REGION Network 2
   // **********************************************************************************************************************
   // 
   // Carrier 81 I-Device Data Transfer Interlocks from Carrier to SDC
   // 
   // **********************************************************************************************************************
   RUNG wire#powerrail
      Coil( "SectionComment" )
   END_RUNG
   // the same network as SCL:
   "SectionComment" := TRUE;
END_REGION

REGION Network 3
   RUNG wire#powerrail
      Contact( "Carrier_81_Status.0" )
      Coil( "EMS".Carrier[81].SDC_IN.HeartBeat )
   END_RUNG
   // the same network as SCL:
   "EMS".Carrier[81].SDC_IN.HeartBeat := "Carrier_81_Status.0";
END_REGION

REGION Network 4
   "C81_Heartbeat_On_Timer".TON(IN := "EMS".Carrier[81].SDC_IN.HeartBeat, PT := T#3s);
END_REGION

REGION Network 5
   "C81_Heartbeat_Off_Timer".TON(IN := NOT "EMS".Carrier[81].SDC_IN.HeartBeat, PT := T#3s);
END_REGION

REGION Network 6
   RUNG wire#powerrail
      Contact( "Carrier_81_Status.7" )
      wire#w1
      Coil( "EMS".Carrier[81].CommFlt )
   END_RUNG
   RUNG wire#powerrail
      Contact( "C81_Heartbeat_On_Timer".Q )
   END_RUNG wire#w1
   RUNG wire#powerrail
      Contact( "C81_Heartbeat_Off_Timer".Q )
   END_RUNG wire#w1
   // the same network as SCL:
   "EMS".Carrier[81].CommFlt := "Carrier_81_Status.7" OR "C81_Heartbeat_On_Timer".Q OR "C81_Heartbeat_Off_Timer".Q;
END_REGION

REGION Network 7
   RUNG wire#powerrail
      Contact( "EMS".Carrier[81].CommFlt )
      JumpCoil( C81_Comm_Fault )
   END_RUNG
   // the same network as SCL:
   IF "EMS".Carrier[81].CommFlt THEN GOTO C81_Comm_Fault; END_IF;
END_REGION

REGION Network 8
   RUNG wire#powerrail
      { S7_Templates := "SrcType := Word" } NE_Contact(in1 := "Carrier_81_CarrierNumber", in2 := 0)
      Move(in := "Carrier_81_CarrierNumber", out1 => "EMS".Carrier[81].SDC_IN.CarrierNumber)
   END_RUNG
   // the same network as SCL:
   IF "Carrier_81_CarrierNumber" <> 0 THEN
       "EMS".Carrier[81].SDC_IN.CarrierNumber := "Carrier_81_CarrierNumber";
   END_IF;
END_REGION

REGION Network 9
   RUNG wire#powerrail
      { S7_Templates := "SrcType := DWord" } NE_Contact(in1 := "Carrier_81_CarrierPosition", in2 := 0)
      Move(in := "Carrier_81_CarrierPosition", out1 => "EMS".Carrier[81].SDC_IN.CarrierPosition)
   END_RUNG
   // the same network as SCL:
   IF "Carrier_81_CarrierPosition" <> 0 THEN
       "EMS".Carrier[81].SDC_IN.CarrierPosition := "Carrier_81_CarrierPosition";
   END_IF;
END_REGION

REGION Network 10
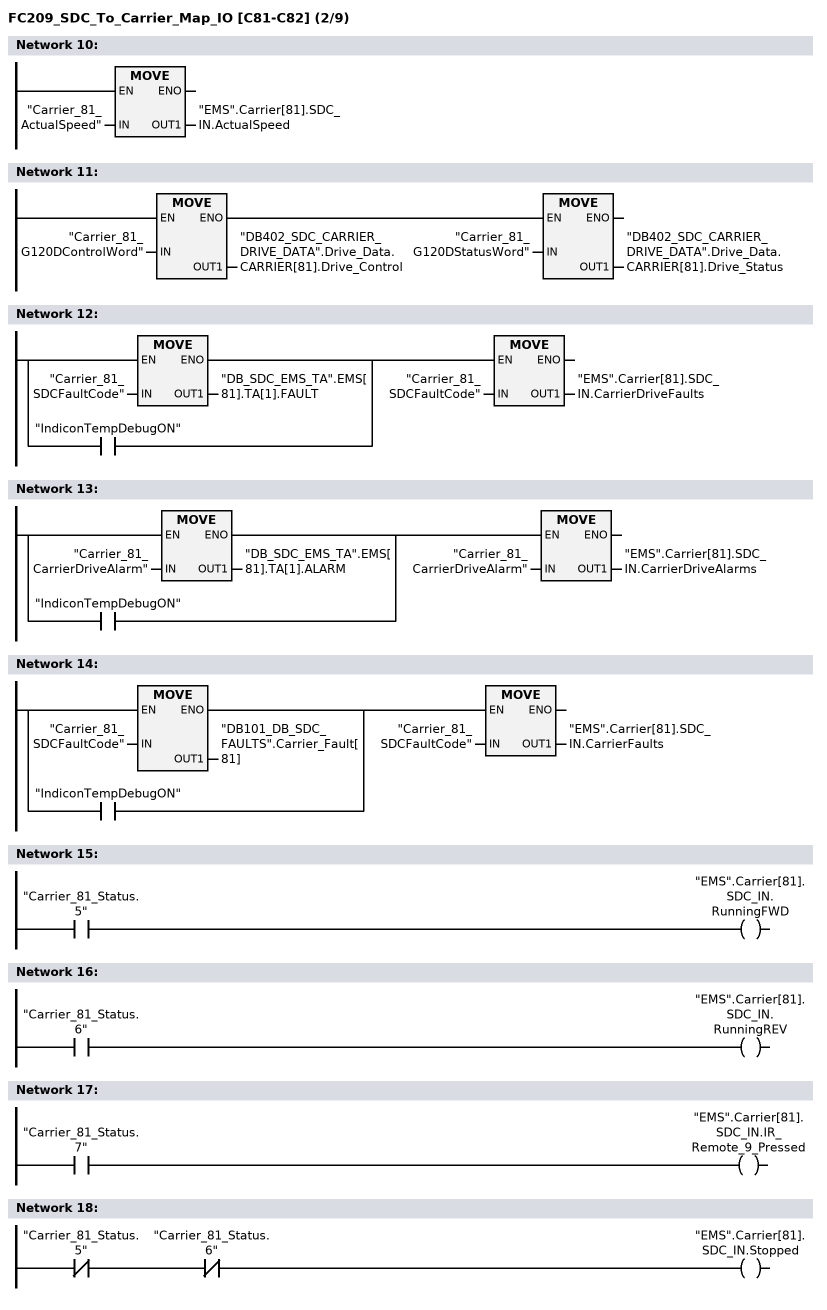
   RUNG wire#powerrail
      Move(in := "Carrier_81_ActualSpeed", out1 => "EMS".Carrier[81].SDC_IN.ActualSpeed)
   END_RUNG
   // the same network as SCL:
   "EMS".Carrier[81].SDC_IN.ActualSpeed := "Carrier_81_ActualSpeed";
END_REGION

REGION Network 11
   RUNG wire#powerrail
      Move(in := "Carrier_81_G120DControlWord", out1 => "DB402_SDC_CARRIER_DRIVE_DATA".Drive_Data.CARRIER[81].Drive_Control)
      Move(in := "Carrier_81_G120DStatusWord", out1 => "DB402_SDC_CARRIER_DRIVE_DATA".Drive_Data.CARRIER[81].Drive_Status)
   END_RUNG
   // the same network as SCL:
   "DB402_SDC_CARRIER_DRIVE_DATA".Drive_Data.CARRIER[81].Drive_Control := "Carrier_81_G120DControlWord";
   "DB402_SDC_CARRIER_DRIVE_DATA".Drive_Data.CARRIER[81].Drive_Status := "Carrier_81_G120DStatusWord";
END_REGION

REGION Network 12
   RUNG wire#powerrail
      Move(in := "Carrier_81_SDCFaultCode", out1 => "DB_SDC_EMS_TA".EMS[81].TA[1].FAULT)
      wire#w1
      Move(in := "Carrier_81_SDCFaultCode", out1 => "EMS".Carrier[81].SDC_IN.CarrierDriveFaults)
   END_RUNG
   RUNG wire#powerrail
      Contact( "IndiconTempDebugON" )
   END_RUNG wire#w1
   // the same network as SCL:
   "DB_SDC_EMS_TA".EMS[81].TA[1].FAULT := "Carrier_81_SDCFaultCode";
   IF TRUE OR "IndiconTempDebugON" THEN
       "EMS".Carrier[81].SDC_IN.CarrierDriveFaults := "Carrier_81_SDCFaultCode";
   END_IF;
END_REGION

REGION Network 13
   RUNG wire#powerrail
      Move(in := "Carrier_81_CarrierDriveAlarm", out1 => "DB_SDC_EMS_TA".EMS[81].TA[1].ALARM)
      wire#w1
      Move(in := "Carrier_81_CarrierDriveAlarm", out1 => "EMS".Carrier[81].SDC_IN.CarrierDriveAlarms)
   END_RUNG
   RUNG wire#powerrail
      Contact( "IndiconTempDebugON" )
   END_RUNG wire#w1
   // the same network as SCL:
   "DB_SDC_EMS_TA".EMS[81].TA[1].ALARM := "Carrier_81_CarrierDriveAlarm";
   IF TRUE OR "IndiconTempDebugON" THEN
       "EMS".Carrier[81].SDC_IN.CarrierDriveAlarms := "Carrier_81_CarrierDriveAlarm";
   END_IF;
END_REGION

REGION Network 14
   RUNG wire#powerrail
      Move(in := "Carrier_81_SDCFaultCode", out1 => "DB101_DB_SDC_FAULTS".Carrier_Fault[81])
      wire#w1
      Move(in := "Carrier_81_SDCFaultCode", out1 => "EMS".Carrier[81].SDC_IN.CarrierFaults)
   END_RUNG
   RUNG wire#powerrail
      Contact( "IndiconTempDebugON" )
   END_RUNG wire#w1
   // the same network as SCL:
   "DB101_DB_SDC_FAULTS".Carrier_Fault[81] := "Carrier_81_SDCFaultCode";
   IF TRUE OR "IndiconTempDebugON" THEN
       "EMS".Carrier[81].SDC_IN.CarrierFaults := "Carrier_81_SDCFaultCode";
   END_IF;
END_REGION

REGION Network 15
   RUNG wire#powerrail
      Contact( "Carrier_81_Status.5" )
      Coil( "EMS".Carrier[81].SDC_IN.RunningFWD )
   END_RUNG
   // the same network as SCL:
   "EMS".Carrier[81].SDC_IN.RunningFWD := "Carrier_81_Status.5";
END_REGION

REGION Network 16
   RUNG wire#powerrail
      Contact( "Carrier_81_Status.6" )
      Coil( "EMS".Carrier[81].SDC_IN.RunningREV )
   END_RUNG
   // the same network as SCL:
   "EMS".Carrier[81].SDC_IN.RunningREV := "Carrier_81_Status.6";
END_REGION

REGION Network 17
   RUNG wire#powerrail
      Contact( "Carrier_81_Status.7" )
      Coil( "EMS".Carrier[81].SDC_IN.IR_Remote_9_Pressed )
   END_RUNG
   // the same network as SCL:
   "EMS".Carrier[81].SDC_IN.IR_Remote_9_Pressed := "Carrier_81_Status.7";
END_REGION

REGION Network 18
   RUNG wire#powerrail
      I_Contact( "Carrier_81_Status.5" )
      I_Contact( "Carrier_81_Status.6" )
      Coil( "EMS".Carrier[81].SDC_IN.Stopped )
   END_RUNG
   // the same network as SCL:
   "EMS".Carrier[81].SDC_IN.Stopped := NOT "Carrier_81_Status.5" AND NOT "Carrier_81_Status.6";
END_REGION

REGION Network 19
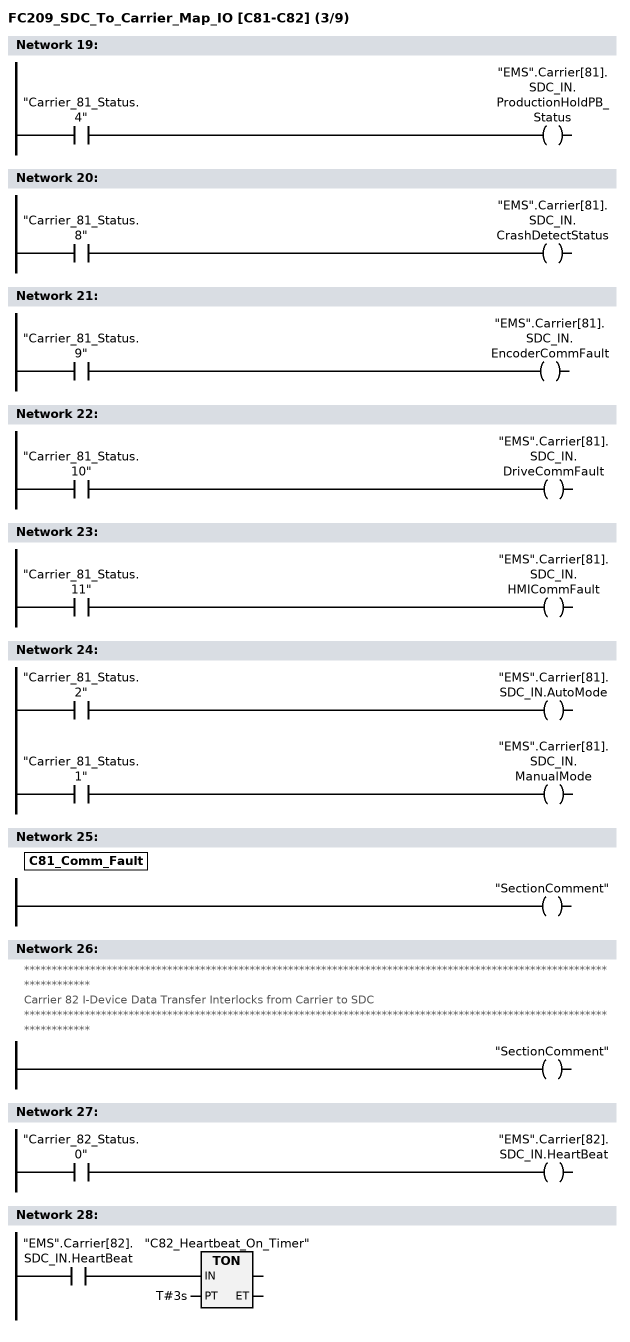
   RUNG wire#powerrail
      Contact( "Carrier_81_Status.4" )
      Coil( "EMS".Carrier[81].SDC_IN.ProductionHoldPB_Status )
   END_RUNG
   // the same network as SCL:
   "EMS".Carrier[81].SDC_IN.ProductionHoldPB_Status := "Carrier_81_Status.4";
END_REGION

REGION Network 20
   RUNG wire#powerrail
      Contact( "Carrier_81_Status.8" )
      Coil( "EMS".Carrier[81].SDC_IN.CrashDetectStatus )
   END_RUNG
   // the same network as SCL:
   "EMS".Carrier[81].SDC_IN.CrashDetectStatus := "Carrier_81_Status.8";
END_REGION

REGION Network 21
   RUNG wire#powerrail
      Contact( "Carrier_81_Status.9" )
      Coil( "EMS".Carrier[81].SDC_IN.EncoderCommFault )
   END_RUNG
   // the same network as SCL:
   "EMS".Carrier[81].SDC_IN.EncoderCommFault := "Carrier_81_Status.9";
END_REGION

REGION Network 22
   RUNG wire#powerrail
      Contact( "Carrier_81_Status.10" )
      Coil( "EMS".Carrier[81].SDC_IN.DriveCommFault )
   END_RUNG
   // the same network as SCL:
   "EMS".Carrier[81].SDC_IN.DriveCommFault := "Carrier_81_Status.10";
END_REGION

REGION Network 23
   RUNG wire#powerrail
      Contact( "Carrier_81_Status.11" )
      Coil( "EMS".Carrier[81].SDC_IN.HMICommFault )
   END_RUNG
   // the same network as SCL:
   "EMS".Carrier[81].SDC_IN.HMICommFault := "Carrier_81_Status.11";
END_REGION

REGION Network 24
   RUNG wire#powerrail
      Contact( "Carrier_81_Status.2" )
      Coil( "EMS".Carrier[81].SDC_IN.AutoMode )
   END_RUNG
   RUNG wire#powerrail
      Contact( "Carrier_81_Status.1" )
      Coil( "EMS".Carrier[81].SDC_IN.ManualMode )
   END_RUNG
   // the same network as SCL:
   "EMS".Carrier[81].SDC_IN.AutoMode := "Carrier_81_Status.2";
   "EMS".Carrier[81].SDC_IN.ManualMode := "Carrier_81_Status.1";
END_REGION

REGION Network 25
   Label( C81_Comm_Fault )
   RUNG wire#powerrail
      Coil( "SectionComment" )
   END_RUNG
   // the same network as SCL:
   C81_Comm_Fault:
   "SectionComment" := TRUE;
END_REGION

REGION Network 26
   // **********************************************************************************************************************
   // 
   // Carrier 82 I-Device Data Transfer Interlocks from Carrier to SDC
   // 
   // **********************************************************************************************************************
   RUNG wire#powerrail
      Coil( "SectionComment" )
   END_RUNG
   // the same network as SCL:
   "SectionComment" := TRUE;
END_REGION

REGION Network 27
   RUNG wire#powerrail
      Contact( "Carrier_82_Status.0" )
      Coil( "EMS".Carrier[82].SDC_IN.HeartBeat )
   END_RUNG
   // the same network as SCL:
   "EMS".Carrier[82].SDC_IN.HeartBeat := "Carrier_82_Status.0";
END_REGION

REGION Network 28
   "C82_Heartbeat_On_Timer".TON(IN := "EMS".Carrier[82].SDC_IN.HeartBeat, PT := T#3s);
END_REGION

REGION Network 29
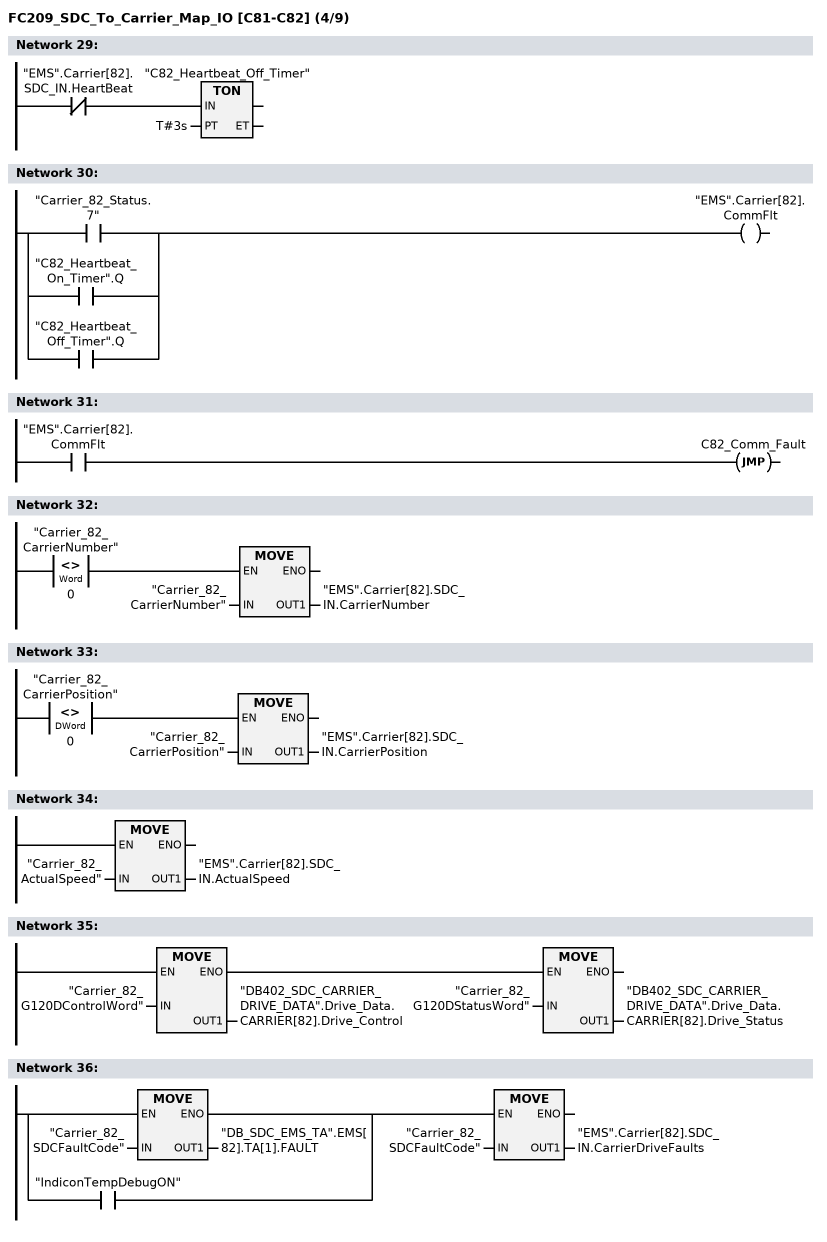
   "C82_Heartbeat_Off_Timer".TON(IN := NOT "EMS".Carrier[82].SDC_IN.HeartBeat, PT := T#3s);
END_REGION

REGION Network 30
   RUNG wire#powerrail
      Contact( "Carrier_82_Status.7" )
      wire#w1
      Coil( "EMS".Carrier[82].CommFlt )
   END_RUNG
   RUNG wire#powerrail
      Contact( "C82_Heartbeat_On_Timer".Q )
   END_RUNG wire#w1
   RUNG wire#powerrail
      Contact( "C82_Heartbeat_Off_Timer".Q )
   END_RUNG wire#w1
   // the same network as SCL:
   "EMS".Carrier[82].CommFlt := "Carrier_82_Status.7" OR "C82_Heartbeat_On_Timer".Q OR "C82_Heartbeat_Off_Timer".Q;
END_REGION

REGION Network 31
   RUNG wire#powerrail
      Contact( "EMS".Carrier[82].CommFlt )
      JumpCoil( C82_Comm_Fault )
   END_RUNG
   // the same network as SCL:
   IF "EMS".Carrier[82].CommFlt THEN GOTO C82_Comm_Fault; END_IF;
END_REGION

REGION Network 32
   RUNG wire#powerrail
      { S7_Templates := "SrcType := Word" } NE_Contact(in1 := "Carrier_82_CarrierNumber", in2 := 0)
      Move(in := "Carrier_82_CarrierNumber", out1 => "EMS".Carrier[82].SDC_IN.CarrierNumber)
   END_RUNG
   // the same network as SCL:
   IF "Carrier_82_CarrierNumber" <> 0 THEN
       "EMS".Carrier[82].SDC_IN.CarrierNumber := "Carrier_82_CarrierNumber";
   END_IF;
END_REGION

REGION Network 33
   RUNG wire#powerrail
      { S7_Templates := "SrcType := DWord" } NE_Contact(in1 := "Carrier_82_CarrierPosition", in2 := 0)
      Move(in := "Carrier_82_CarrierPosition", out1 => "EMS".Carrier[82].SDC_IN.CarrierPosition)
   END_RUNG
   // the same network as SCL:
   IF "Carrier_82_CarrierPosition" <> 0 THEN
       "EMS".Carrier[82].SDC_IN.CarrierPosition := "Carrier_82_CarrierPosition";
   END_IF;
END_REGION

REGION Network 34
   RUNG wire#powerrail
      Move(in := "Carrier_82_ActualSpeed", out1 => "EMS".Carrier[82].SDC_IN.ActualSpeed)
   END_RUNG
   // the same network as SCL:
   "EMS".Carrier[82].SDC_IN.ActualSpeed := "Carrier_82_ActualSpeed";
END_REGION

REGION Network 35
   RUNG wire#powerrail
      Move(in := "Carrier_82_G120DControlWord", out1 => "DB402_SDC_CARRIER_DRIVE_DATA".Drive_Data.CARRIER[82].Drive_Control)
      Move(in := "Carrier_82_G120DStatusWord", out1 => "DB402_SDC_CARRIER_DRIVE_DATA".Drive_Data.CARRIER[82].Drive_Status)
   END_RUNG
   // the same network as SCL:
   "DB402_SDC_CARRIER_DRIVE_DATA".Drive_Data.CARRIER[82].Drive_Control := "Carrier_82_G120DControlWord";
   "DB402_SDC_CARRIER_DRIVE_DATA".Drive_Data.CARRIER[82].Drive_Status := "Carrier_82_G120DStatusWord";
END_REGION

REGION Network 36
   RUNG wire#powerrail
      Move(in := "Carrier_82_SDCFaultCode", out1 => "DB_SDC_EMS_TA".EMS[82].TA[1].FAULT)
      wire#w1
      Move(in := "Carrier_82_SDCFaultCode", out1 => "EMS".Carrier[82].SDC_IN.CarrierDriveFaults)
   END_RUNG
   RUNG wire#powerrail
      Contact( "IndiconTempDebugON" )
   END_RUNG wire#w1
   // the same network as SCL:
   "DB_SDC_EMS_TA".EMS[82].TA[1].FAULT := "Carrier_82_SDCFaultCode";
   IF TRUE OR "IndiconTempDebugON" THEN
       "EMS".Carrier[82].SDC_IN.CarrierDriveFaults := "Carrier_82_SDCFaultCode";
   END_IF;
END_REGION

REGION Network 37
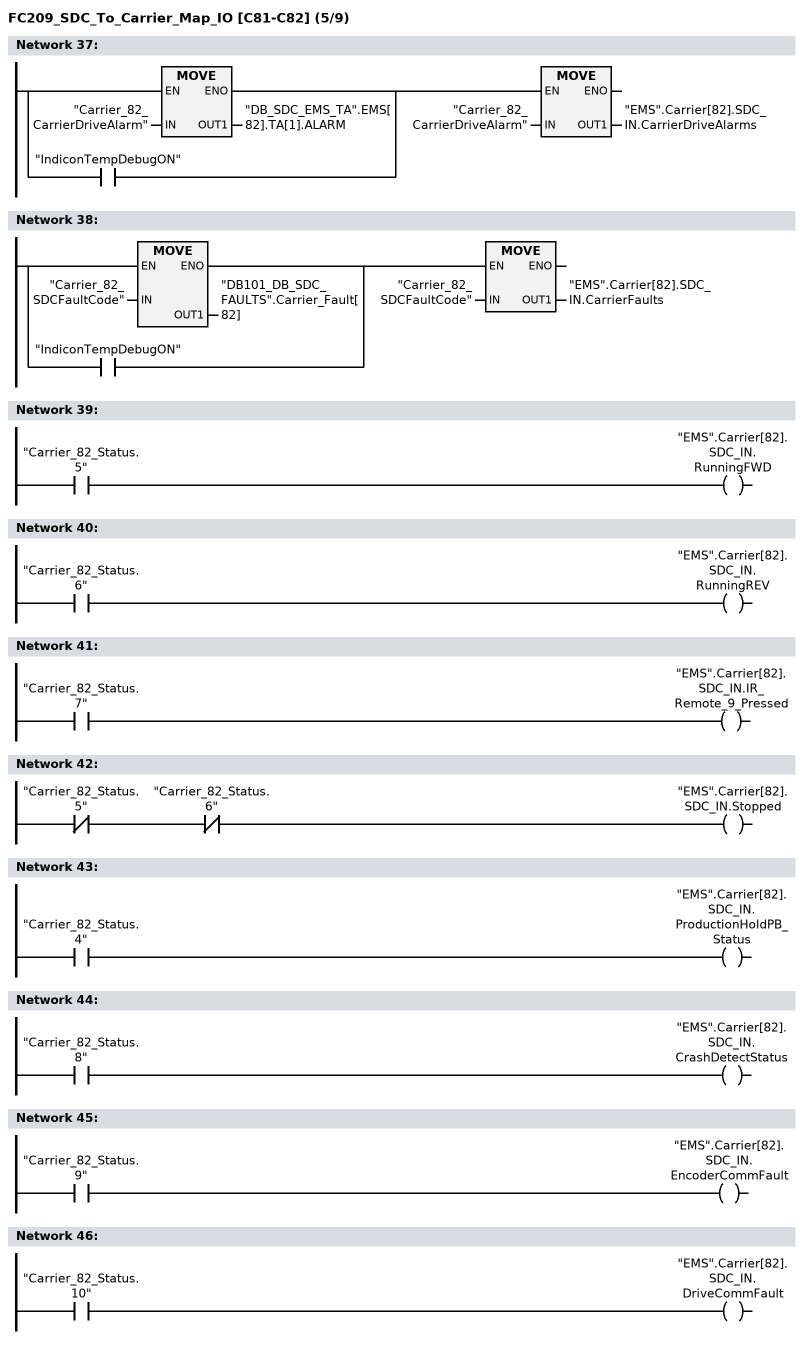
   RUNG wire#powerrail
      Move(in := "Carrier_82_CarrierDriveAlarm", out1 => "DB_SDC_EMS_TA".EMS[82].TA[1].ALARM)
      wire#w1
      Move(in := "Carrier_82_CarrierDriveAlarm", out1 => "EMS".Carrier[82].SDC_IN.CarrierDriveAlarms)
   END_RUNG
   RUNG wire#powerrail
      Contact( "IndiconTempDebugON" )
   END_RUNG wire#w1
   // the same network as SCL:
   "DB_SDC_EMS_TA".EMS[82].TA[1].ALARM := "Carrier_82_CarrierDriveAlarm";
   IF TRUE OR "IndiconTempDebugON" THEN
       "EMS".Carrier[82].SDC_IN.CarrierDriveAlarms := "Carrier_82_CarrierDriveAlarm";
   END_IF;
END_REGION

REGION Network 38
   RUNG wire#powerrail
      Move(in := "Carrier_82_SDCFaultCode", out1 => "DB101_DB_SDC_FAULTS".Carrier_Fault[82])
      wire#w1
      Move(in := "Carrier_82_SDCFaultCode", out1 => "EMS".Carrier[82].SDC_IN.CarrierFaults)
   END_RUNG
   RUNG wire#powerrail
      Contact( "IndiconTempDebugON" )
   END_RUNG wire#w1
   // the same network as SCL:
   "DB101_DB_SDC_FAULTS".Carrier_Fault[82] := "Carrier_82_SDCFaultCode";
   IF TRUE OR "IndiconTempDebugON" THEN
       "EMS".Carrier[82].SDC_IN.CarrierFaults := "Carrier_82_SDCFaultCode";
   END_IF;
END_REGION

REGION Network 39
   RUNG wire#powerrail
      Contact( "Carrier_82_Status.5" )
      Coil( "EMS".Carrier[82].SDC_IN.RunningFWD )
   END_RUNG
   // the same network as SCL:
   "EMS".Carrier[82].SDC_IN.RunningFWD := "Carrier_82_Status.5";
END_REGION

REGION Network 40
   RUNG wire#powerrail
      Contact( "Carrier_82_Status.6" )
      Coil( "EMS".Carrier[82].SDC_IN.RunningREV )
   END_RUNG
   // the same network as SCL:
   "EMS".Carrier[82].SDC_IN.RunningREV := "Carrier_82_Status.6";
END_REGION

REGION Network 41
   RUNG wire#powerrail
      Contact( "Carrier_82_Status.7" )
      Coil( "EMS".Carrier[82].SDC_IN.IR_Remote_9_Pressed )
   END_RUNG
   // the same network as SCL:
   "EMS".Carrier[82].SDC_IN.IR_Remote_9_Pressed := "Carrier_82_Status.7";
END_REGION

REGION Network 42
   RUNG wire#powerrail
      I_Contact( "Carrier_82_Status.5" )
      I_Contact( "Carrier_82_Status.6" )
      Coil( "EMS".Carrier[82].SDC_IN.Stopped )
   END_RUNG
   // the same network as SCL:
   "EMS".Carrier[82].SDC_IN.Stopped := NOT "Carrier_82_Status.5" AND NOT "Carrier_82_Status.6";
END_REGION

REGION Network 43
   RUNG wire#powerrail
      Contact( "Carrier_82_Status.4" )
      Coil( "EMS".Carrier[82].SDC_IN.ProductionHoldPB_Status )
   END_RUNG
   // the same network as SCL:
   "EMS".Carrier[82].SDC_IN.ProductionHoldPB_Status := "Carrier_82_Status.4";
END_REGION

REGION Network 44
   RUNG wire#powerrail
      Contact( "Carrier_82_Status.8" )
      Coil( "EMS".Carrier[82].SDC_IN.CrashDetectStatus )
   END_RUNG
   // the same network as SCL:
   "EMS".Carrier[82].SDC_IN.CrashDetectStatus := "Carrier_82_Status.8";
END_REGION

REGION Network 45
   RUNG wire#powerrail
      Contact( "Carrier_82_Status.9" )
      Coil( "EMS".Carrier[82].SDC_IN.EncoderCommFault )
   END_RUNG
   // the same network as SCL:
   "EMS".Carrier[82].SDC_IN.EncoderCommFault := "Carrier_82_Status.9";
END_REGION

REGION Network 46
   RUNG wire#powerrail
      Contact( "Carrier_82_Status.10" )
      Coil( "EMS".Carrier[82].SDC_IN.DriveCommFault )
   END_RUNG
   // the same network as SCL:
   "EMS".Carrier[82].SDC_IN.DriveCommFault := "Carrier_82_Status.10";
END_REGION

REGION Network 47
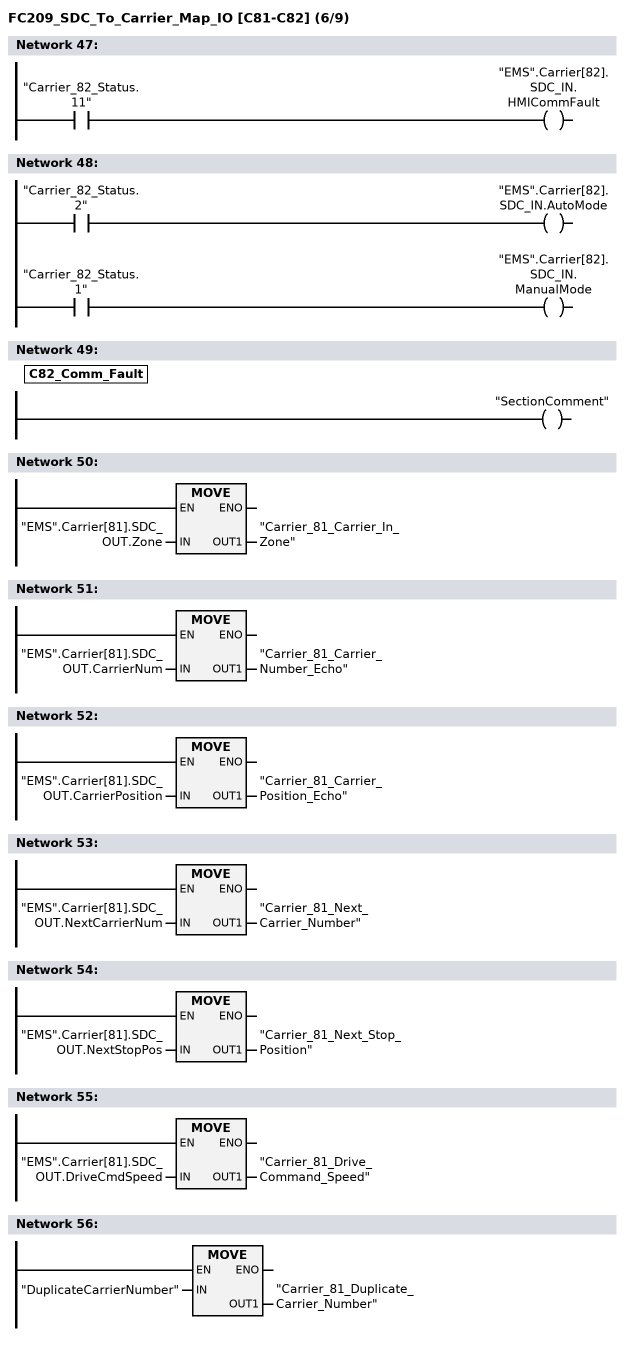
   RUNG wire#powerrail
      Contact( "Carrier_82_Status.11" )
      Coil( "EMS".Carrier[82].SDC_IN.HMICommFault )
   END_RUNG
   // the same network as SCL:
   "EMS".Carrier[82].SDC_IN.HMICommFault := "Carrier_82_Status.11";
END_REGION

REGION Network 48
   RUNG wire#powerrail
      Contact( "Carrier_82_Status.2" )
      Coil( "EMS".Carrier[82].SDC_IN.AutoMode )
   END_RUNG
   RUNG wire#powerrail
      Contact( "Carrier_82_Status.1" )
      Coil( "EMS".Carrier[82].SDC_IN.ManualMode )
   END_RUNG
   // the same network as SCL:
   "EMS".Carrier[82].SDC_IN.AutoMode := "Carrier_82_Status.2";
   "EMS".Carrier[82].SDC_IN.ManualMode := "Carrier_82_Status.1";
END_REGION

REGION Network 49
   Label( C82_Comm_Fault )
   RUNG wire#powerrail
      Coil( "SectionComment" )
   END_RUNG
   // the same network as SCL:
   C82_Comm_Fault:
   "SectionComment" := TRUE;
END_REGION

REGION Network 50
   RUNG wire#powerrail
      Move(in := "EMS".Carrier[81].SDC_OUT.Zone, out1 => "Carrier_81_Carrier_In_Zone")
   END_RUNG
   // the same network as SCL:
   "Carrier_81_Carrier_In_Zone" := "EMS".Carrier[81].SDC_OUT.Zone;
END_REGION

REGION Network 51
   RUNG wire#powerrail
      Move(in := "EMS".Carrier[81].SDC_OUT.CarrierNum, out1 => "Carrier_81_Carrier_Number_Echo")
   END_RUNG
   // the same network as SCL:
   "Carrier_81_Carrier_Number_Echo" := "EMS".Carrier[81].SDC_OUT.CarrierNum;
END_REGION

REGION Network 52
   RUNG wire#powerrail
      Move(in := "EMS".Carrier[81].SDC_OUT.CarrierPosition, out1 => "Carrier_81_Carrier_Position_Echo")
   END_RUNG
   // the same network as SCL:
   "Carrier_81_Carrier_Position_Echo" := "EMS".Carrier[81].SDC_OUT.CarrierPosition;
END_REGION

REGION Network 53
   RUNG wire#powerrail
      Move(in := "EMS".Carrier[81].SDC_OUT.NextCarrierNum, out1 => "Carrier_81_Next_Carrier_Number")
   END_RUNG
   // the same network as SCL:
   "Carrier_81_Next_Carrier_Number" := "EMS".Carrier[81].SDC_OUT.NextCarrierNum;
END_REGION

REGION Network 54
   RUNG wire#powerrail
      Move(in := "EMS".Carrier[81].SDC_OUT.NextStopPos, out1 => "Carrier_81_Next_Stop_Position")
   END_RUNG
   // the same network as SCL:
   "Carrier_81_Next_Stop_Position" := "EMS".Carrier[81].SDC_OUT.NextStopPos;
END_REGION

REGION Network 55
   RUNG wire#powerrail
      Move(in := "EMS".Carrier[81].SDC_OUT.DriveCmdSpeed, out1 => "Carrier_81_Drive_Command_Speed")
   END_RUNG
   // the same network as SCL:
   "Carrier_81_Drive_Command_Speed" := "EMS".Carrier[81].SDC_OUT.DriveCmdSpeed;
END_REGION

REGION Network 56
   RUNG wire#powerrail
      Move(in := "DuplicateCarrierNumber", out1 => "Carrier_81_Duplicate_Carrier_Number")
   END_RUNG
   // the same network as SCL:
   "Carrier_81_Duplicate_Carrier_Number" := "DuplicateCarrierNumber";
END_REGION

REGION Network 57
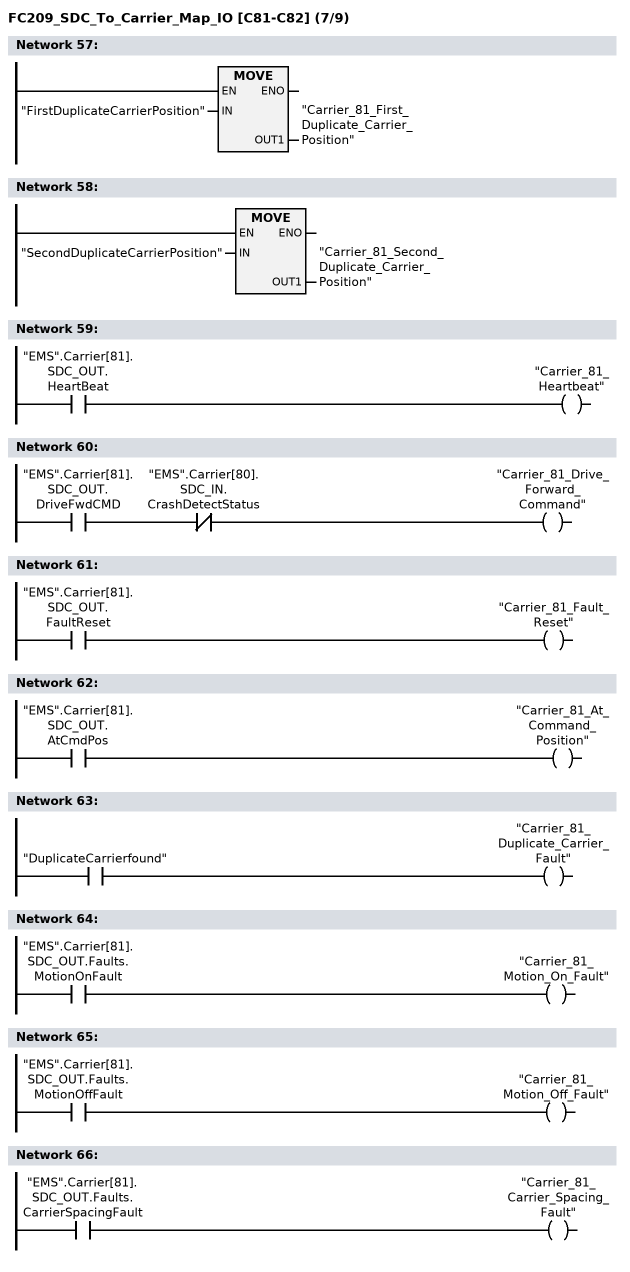
   RUNG wire#powerrail
      Move(in := "FirstDuplicateCarrierPosition", out1 => "Carrier_81_First_Duplicate_Carrier_Position")
   END_RUNG
   // the same network as SCL:
   "Carrier_81_First_Duplicate_Carrier_Position" := "FirstDuplicateCarrierPosition";
END_REGION

REGION Network 58
   RUNG wire#powerrail
      Move(in := "SecondDuplicateCarrierPosition", out1 => "Carrier_81_Second_Duplicate_Carrier_Position")
   END_RUNG
   // the same network as SCL:
   "Carrier_81_Second_Duplicate_Carrier_Position" := "SecondDuplicateCarrierPosition";
END_REGION

REGION Network 59
   RUNG wire#powerrail
      Contact( "EMS".Carrier[81].SDC_OUT.HeartBeat )
      Coil( "Carrier_81_Heartbeat" )
   END_RUNG
   // the same network as SCL:
   "Carrier_81_Heartbeat" := "EMS".Carrier[81].SDC_OUT.HeartBeat;
END_REGION

REGION Network 60
   RUNG wire#powerrail
      Contact( "EMS".Carrier[81].SDC_OUT.DriveFwdCMD )
      I_Contact( "EMS".Carrier[80].SDC_IN.CrashDetectStatus )
      Coil( "Carrier_81_Drive_Forward_Command" )
   END_RUNG
   // the same network as SCL:
   "Carrier_81_Drive_Forward_Command" := "EMS".Carrier[81].SDC_OUT.DriveFwdCMD AND NOT "EMS".Carrier[80].SDC_IN.CrashDetectStatus;
END_REGION

REGION Network 61
   RUNG wire#powerrail
      Contact( "EMS".Carrier[81].SDC_OUT.FaultReset )
      Coil( "Carrier_81_Fault_Reset" )
   END_RUNG
   // the same network as SCL:
   "Carrier_81_Fault_Reset" := "EMS".Carrier[81].SDC_OUT.FaultReset;
END_REGION

REGION Network 62
   RUNG wire#powerrail
      Contact( "EMS".Carrier[81].SDC_OUT.AtCmdPos )
      Coil( "Carrier_81_At_Command_Position" )
   END_RUNG
   // the same network as SCL:
   "Carrier_81_At_Command_Position" := "EMS".Carrier[81].SDC_OUT.AtCmdPos;
END_REGION

REGION Network 63
   RUNG wire#powerrail
      Contact( "DuplicateCarrierfound" )
      Coil( "Carrier_81_Duplicate_Carrier_Fault" )
   END_RUNG
   // the same network as SCL:
   "Carrier_81_Duplicate_Carrier_Fault" := "DuplicateCarrierfound";
END_REGION

REGION Network 64
   RUNG wire#powerrail
      Contact( "EMS".Carrier[81].SDC_OUT.Faults.MotionOnFault )
      Coil( "Carrier_81_Motion_On_Fault" )
   END_RUNG
   // the same network as SCL:
   "Carrier_81_Motion_On_Fault" := "EMS".Carrier[81].SDC_OUT.Faults.MotionOnFault;
END_REGION

REGION Network 65
   RUNG wire#powerrail
      Contact( "EMS".Carrier[81].SDC_OUT.Faults.MotionOffFault )
      Coil( "Carrier_81_Motion_Off_Fault" )
   END_RUNG
   // the same network as SCL:
   "Carrier_81_Motion_Off_Fault" := "EMS".Carrier[81].SDC_OUT.Faults.MotionOffFault;
END_REGION

REGION Network 66
   RUNG wire#powerrail
      Contact( "EMS".Carrier[81].SDC_OUT.Faults.CarrierSpacingFault )
      Coil( "Carrier_81_Carrier_Spacing_Fault" )
   END_RUNG
   // the same network as SCL:
   "Carrier_81_Carrier_Spacing_Fault" := "EMS".Carrier[81].SDC_OUT.Faults.CarrierSpacingFault;
END_REGION

REGION Network 67
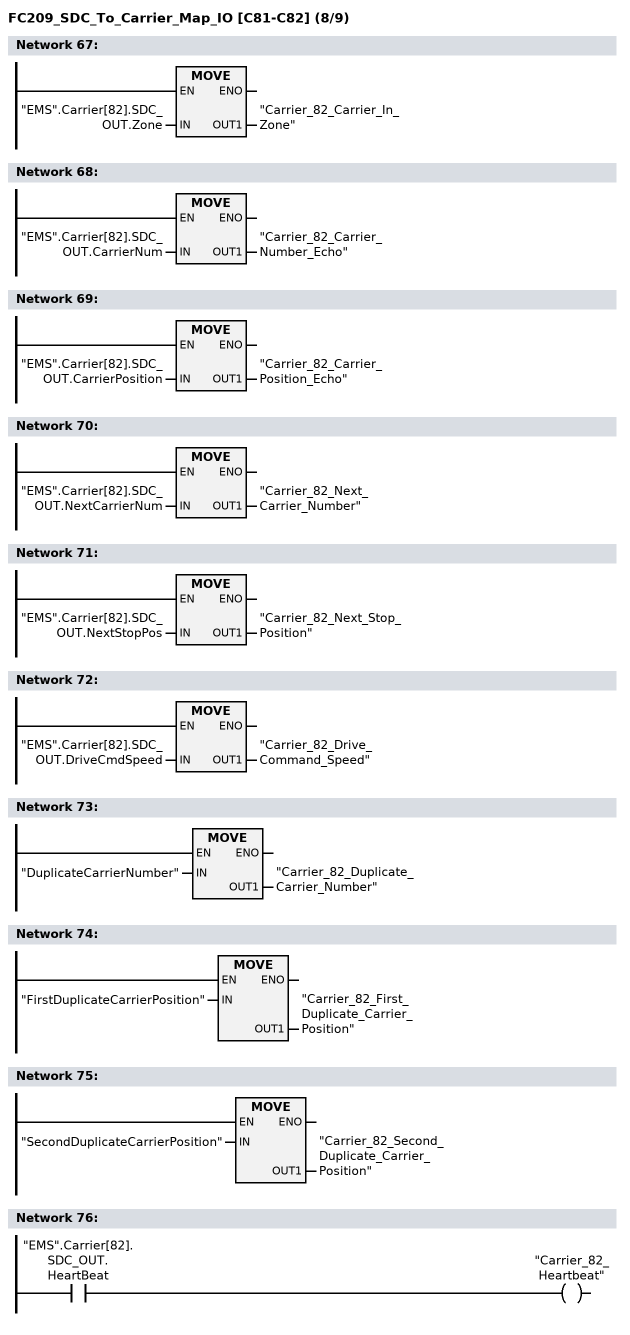
   RUNG wire#powerrail
      Move(in := "EMS".Carrier[82].SDC_OUT.Zone, out1 => "Carrier_82_Carrier_In_Zone")
   END_RUNG
   // the same network as SCL:
   "Carrier_82_Carrier_In_Zone" := "EMS".Carrier[82].SDC_OUT.Zone;
END_REGION

REGION Network 68
   RUNG wire#powerrail
      Move(in := "EMS".Carrier[82].SDC_OUT.CarrierNum, out1 => "Carrier_82_Carrier_Number_Echo")
   END_RUNG
   // the same network as SCL:
   "Carrier_82_Carrier_Number_Echo" := "EMS".Carrier[82].SDC_OUT.CarrierNum;
END_REGION

REGION Network 69
   RUNG wire#powerrail
      Move(in := "EMS".Carrier[82].SDC_OUT.CarrierPosition, out1 => "Carrier_82_Carrier_Position_Echo")
   END_RUNG
   // the same network as SCL:
   "Carrier_82_Carrier_Position_Echo" := "EMS".Carrier[82].SDC_OUT.CarrierPosition;
END_REGION

REGION Network 70
   RUNG wire#powerrail
      Move(in := "EMS".Carrier[82].SDC_OUT.NextCarrierNum, out1 => "Carrier_82_Next_Carrier_Number")
   END_RUNG
   // the same network as SCL:
   "Carrier_82_Next_Carrier_Number" := "EMS".Carrier[82].SDC_OUT.NextCarrierNum;
END_REGION

REGION Network 71
   RUNG wire#powerrail
      Move(in := "EMS".Carrier[82].SDC_OUT.NextStopPos, out1 => "Carrier_82_Next_Stop_Position")
   END_RUNG
   // the same network as SCL:
   "Carrier_82_Next_Stop_Position" := "EMS".Carrier[82].SDC_OUT.NextStopPos;
END_REGION

REGION Network 72
   RUNG wire#powerrail
      Move(in := "EMS".Carrier[82].SDC_OUT.DriveCmdSpeed, out1 => "Carrier_82_Drive_Command_Speed")
   END_RUNG
   // the same network as SCL:
   "Carrier_82_Drive_Command_Speed" := "EMS".Carrier[82].SDC_OUT.DriveCmdSpeed;
END_REGION

REGION Network 73
   RUNG wire#powerrail
      Move(in := "DuplicateCarrierNumber", out1 => "Carrier_82_Duplicate_Carrier_Number")
   END_RUNG
   // the same network as SCL:
   "Carrier_82_Duplicate_Carrier_Number" := "DuplicateCarrierNumber";
END_REGION

REGION Network 74
   RUNG wire#powerrail
      Move(in := "FirstDuplicateCarrierPosition", out1 => "Carrier_82_First_Duplicate_Carrier_Position")
   END_RUNG
   // the same network as SCL:
   "Carrier_82_First_Duplicate_Carrier_Position" := "FirstDuplicateCarrierPosition";
END_REGION

REGION Network 75
   RUNG wire#powerrail
      Move(in := "SecondDuplicateCarrierPosition", out1 => "Carrier_82_Second_Duplicate_Carrier_Position")
   END_RUNG
   // the same network as SCL:
   "Carrier_82_Second_Duplicate_Carrier_Position" := "SecondDuplicateCarrierPosition";
END_REGION

REGION Network 76
   RUNG wire#powerrail
      Contact( "EMS".Carrier[82].SDC_OUT.HeartBeat )
      Coil( "Carrier_82_Heartbeat" )
   END_RUNG
   // the same network as SCL:
   "Carrier_82_Heartbeat" := "EMS".Carrier[82].SDC_OUT.HeartBeat;
END_REGION

REGION Network 77
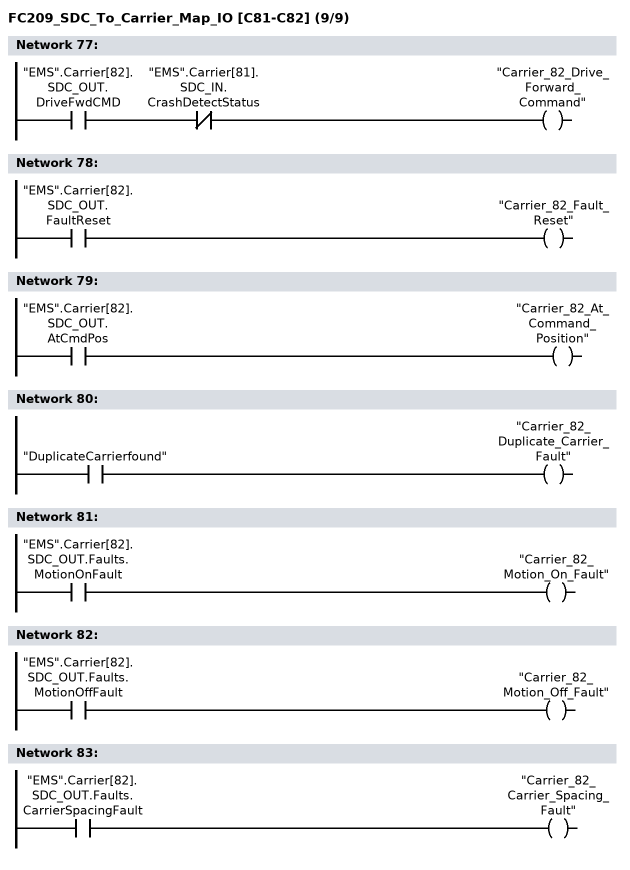
   RUNG wire#powerrail
      Contact( "EMS".Carrier[82].SDC_OUT.DriveFwdCMD )
      I_Contact( "EMS".Carrier[81].SDC_IN.CrashDetectStatus )
      Coil( "Carrier_82_Drive_Forward_Command" )
   END_RUNG
   // the same network as SCL:
   "Carrier_82_Drive_Forward_Command" := "EMS".Carrier[82].SDC_OUT.DriveFwdCMD AND NOT "EMS".Carrier[81].SDC_IN.CrashDetectStatus;
END_REGION

REGION Network 78
   RUNG wire#powerrail
      Contact( "EMS".Carrier[82].SDC_OUT.FaultReset )
      Coil( "Carrier_82_Fault_Reset" )
   END_RUNG
   // the same network as SCL:
   "Carrier_82_Fault_Reset" := "EMS".Carrier[82].SDC_OUT.FaultReset;
END_REGION

REGION Network 79
   RUNG wire#powerrail
      Contact( "EMS".Carrier[82].SDC_OUT.AtCmdPos )
      Coil( "Carrier_82_At_Command_Position" )
   END_RUNG
   // the same network as SCL:
   "Carrier_82_At_Command_Position" := "EMS".Carrier[82].SDC_OUT.AtCmdPos;
END_REGION
